// TIA Portal project "PolyMix_v0.1" (V14)

(* hardware
DEVICE "S7-1200 station_1"  S7-1200 Station
   slot 0: "Rack_0"  S7-1200 Rack  Rack  V1.0
   slot 1: "PLC_PolyMix_001"  CPU 1214C DC/DC/DC  6ES7 214-1AG40-0XB0  V4.2
DEVICE "HMI_PolyMix_001"  KTP700 Basic PN
   slot 0: "KTP700 Basic PN"  KTP700 Basic PN  6AV2 123-2GB03-0AX0  14.0.1.0
   slot 1: "HMI_RT_1"  KTP700 Basic PN  6AV2 123-2GB03-0AX0  14.0.1.0
   slot 5: "HMI_PolyMix_001.IE_CP_1"  PROFINET Interface  14.0.1.0
      slot 1: "PROFINET Interface_1"  PROFINET Interface
         slot 1: "Port_1"  Port
DEVICE "S7-1200 station_2"  S7-1200 Station
   slot 0: "Rack_0"  S7-1200 Rack  Rack  V1.0
   slot 1: "PLC_Master"  CPU 1214C DC/DC/DC  6ES7 214-1AG40-0XB0  V4.2
   slot 2: "AI 4x13BIT/AQ 2x14BIT_1"  6ES7 234-4HE32-0XB0  V2.0
   slot 3: "AI 4x13BIT/AQ 2x14BIT_2"  6ES7 234-4HE32-0XB0  V2.0
   slot 101: "CM 1241 (RS232)_1"  6ES7 241-1AH32-0XB0  V2.2
   slot 102: "CM 1241 (RS232)_2"  6ES7 241-1AH32-0XB0  V2.2
DEVICE "S7-1200 station_3"  S7-1200 Station
   slot 0: "Rack_0"  S7-1200 Rack  Rack  V1.0
   slot 1: "PLC_PolyMix_002"  CPU 1214C DC/DC/DC  6ES7 214-1AG40-0XB0  V4.2
DEVICE "HMI_PolyMix_002"  KTP700 Basic PN
   slot 0: "KTP700 Basic PN"  KTP700 Basic PN  6AV2 123-2GB03-0AX0  14.0.1.0
   slot 1: "HMI_RT_2"  KTP700 Basic PN  6AV2 123-2GB03-0AX0  14.0.1.0
   slot 5: "HMI_PolyMix_002.1.IE_CP_1"  PROFINET Interface  14.0.1.0
      slot 1: "PROFINET Interface_1"  PROFINET Interface
         slot 1: "Port_1"  Port
DEVICE "HMI_Master"  KTP700 Basic PN
   slot 0: "KTP700 Basic PN"  KTP700 Basic PN  6AV2 123-2GB03-0AX0  14.0.1.0
   slot 1: "HMI_RT_3"  KTP700 Basic PN  6AV2 123-2GB03-0AX0  14.0.1.0
   slot 5: "HMI_Master.2.1.IE_CP_1"  PROFINET Interface  14.0.1.0
      slot 1: "PROFINET Interface_1"  PROFINET Interface
         slot 1: "Port_1"  Port
DEVICE "HMI_Master_1"  KTP700 Basic PN
   slot 0: "KTP700 Basic PN"  KTP700 Basic PN  6AV2 123-2GB03-0AX0  14.0.1.0
   slot 1: "HMI_RT_4"  KTP700 Basic PN  6AV2 123-2GB03-0AX0  14.0.1.0
   slot 5: "HMI_Master.2.1.IE_CP_1"  PROFINET Interface  14.0.1.0
      slot 1: "PROFINET Interface_1"  PROFINET Interface
         slot 1: "Port_1"  Port
*)

// ===== PLC "PLC_PolyMix_001"  CPU 1214C DC/DC/DC =====
// protected blocks, not shown: "AI_ex", "AIx", "AO_ex", "DRV_M_D", "FlowMeter", "Logick", "Motors", "PLF_FC", "Time_m", "Time_r", "Time_s"

VAR_GLOBAL   // PLC tag table "Default tag table"
   "Mix_1_Clock" AT %M10.0 : Bool;
   "Mix_2_Clock" AT %M10.1 : Bool;
   "Mix_3_Clock" AT %M10.2 : Bool;
   "Flow" AT %IW256 : Int;
   "Level" AT %IW258 : Int;
END_VAR

VAR_GLOBAL   // PLC tag table "Sys"
   "pulse_01s" AT %M2.0 : Bool;
   "pulse_05s" AT %M2.1 : Bool;
   "pulse_1s" AT %M2.2 : Bool;
   "All_block" AT %M3.0 : Bool;
   "Reset_All" AT %M3.1 : Bool;
   "Sim_All" AT %M3.2 : Bool;
   "Any_Hand" AT %M5.0 : Bool;
   "DI_Hand" AT %M5.1 : Bool;
   "DO_Hand" AT %M5.2 : Bool;
   "AI_Hand" AT %M5.3 : Bool;
   "AO_Hand" AT %M5.4 : Bool;
   "M_Hand" AT %M5.5 : Bool;
   "V_Hand" AT %M5.6 : Bool;
   "X_Hand" AT %M5.7 : Bool;
   "System_Byte" AT %MB1 : Byte;
   "FirstScan" AT %M1.0 : Bool;
   "DiagStatusUpdate" AT %M1.1 : Bool;
   "ON" AT %M1.2 : Bool;
   "OFF" AT %M1.3 : Bool;
   "Clock_Byte" AT %MB0 : Byte;
   "Clock_10Hz" AT %M0.0 : Bool;
   "Clock_5Hz" AT %M0.1 : Bool;
   "Clock_2.5Hz" AT %M0.2 : Bool;
   "Clock_2Hz" AT %M0.3 : Bool;
   "Clock_1.25Hz" AT %M0.4 : Bool;
   "Clock_1Hz" AT %M0.5 : Bool;
   "Clock_0.625Hz" AT %M0.6 : Bool;
   "Clock_0.5Hz" AT %M0.7 : Bool;
   "F_pulse_01s" AT %M2.3 : Bool;
   "F_pulse_05s" AT %M2.4 : Bool;
   "F_pulse_1s" AT %M2.5 : Bool;
   "FN_pulse_01s" AT %M2.6 : Bool;
   "Clock_5s" AT %M2.7 : Bool;
   "Any_Alm" AT %M6.0 : Bool;
   "AI_Alm" AT %M6.1 : Bool;
   "M_Alm" AT %M6.2 : Bool;
   "V_Alm" AT %M6.3 : Bool;
   "C_Alm" AT %M6.4 : Bool;
   "N_Alm" AT %M6.5 : Bool;
   "L_Alm" AT %M6.6 : Bool;
   "X_Alm" AT %M6.7 : Bool;
END_VAR

VAR_GLOBAL   // PLC tag table "IO Table"
   "DD_FB_Ready" AT %I0.6 : Bool;   // I 0.6 - Дозатор сухого вещества - готовность
   "Dos_FB_Run" AT %I0.7 : Bool;   // I 0.7 - Дозатор - работа
   "DD_LLS" AT %I1.0 : Bool;   // I 1.0 - Дозатор сухого вещества - низкий уровень
   "Vibro_FB_Ready" AT %I1.1 : Bool;   // I 1.1 - Вибратор - готовность
   "Transporter" AT %I1.2 : Bool;   // I 1.2 - Пневмотранспортёр - готовность
   "DL_FB_Ready" AT %I1.3 : Bool;   // I 1.3 - Дозатор жидкого вещества - готовность
   "Dry_Run" AT %I1.4 : Bool;   // I 1.4 - Датчик протока
   "AllBlock" AT %I1.5 : Bool;   // I 1.5 - Датчик перелива или Аварийная остановка
   "M1_FB_Ready" AT %I0.0 : Bool;   // I 0.0 - Мешалка 1 - готовность
   "M1_FB_Run" AT %I0.1 : Bool;   // I 0.1 - Мешалка 1 - работа
   "M2_FB_Ready" AT %I0.2 : Bool;   // I 0.2 - Мешалка 2 - готовность
   "M2_FB_Run" AT %I0.3 : Bool;   // I 0.3 - Мешалка 2 - работа
   "M3_FB_Ready" AT %I0.4 : Bool;   // I 0.4 - Мешалка 3 - готовность
   "M3_FB_Run" AT %I0.5 : Bool;   // I 0.5 - Мешалка 3 - работа
   "M1_CMD" AT %Q0.0 : Bool;   // Q 0.0 - Мешалка 1 - запуск
   "M2_CMD" AT %Q0.1 : Bool;   // Q 0.1 - Мешалка 2 - запуск
   "M3_CMD" AT %Q0.2 : Bool;   // Q 0.2 - Мешалка 3 - запуск
   "DD_CMD" AT %Q0.3 : Bool;   // Q 0.3 - Дозатор сухого вещества - запуск
   "Vibro_CMD" AT %Q0.4 : Bool;   // Q 0.4 - Вибратор - запуск
   "DL_CMD" AT %Q0.5 : Bool;   // Q 0.5 - Дозатор жидкого вещества - запуск
   "KC1_CMD" AT %Q0.6 : Bool;   // Q 0.6 - Соленоидный клапан КС1
   "LED_Dry_Run" AT %Q0.7 : Bool;   // Q 0.7 - LED - сухой ход
   "LED_Alarm" AT %Q1.0 : Bool;   // Q 1.0 - LED - общая авария
   "LED_Empty" AT %Q1.1 : Bool;   // Q 1.1 - LED - бункер пуст
END_VAR

DATA_BLOCK "Any_DB"   // DB3
{ S7_Optimized_Access := 'FALSE' }
VERSION : 0.1
   VAR
      Level_M : Int;
      Level_S : Int;
      Flow_M : Int;
      Flow_S : Int;
      DD_View : Bool;
      Level_View : Bool;
   END_VAR
BEGIN
END_DATA_BLOCK

DATA_BLOCK "CONFIG"   // DB10
{ S7_Optimized_Access := 'FALSE' }
VERSION : 0.1
   VAR
      Config : Struct
         Use_DD : Bool;   // Использовать сухой дозатор
         Use_DL : Bool := true;   // Использовать жидкий дозатор
         Use_Mix_1 : Bool := true;   // Использовать мешалку 1
         Use_Mix_2 : Bool := true;   // Использовать мешалку 2
         Use_Mix_3 : Bool := true;   // Использовать мешалку 3
      END_STRUCT;
   END_VAR
BEGIN
END_DATA_BLOCK

DATA_BLOCK "Comm_DB"   // DB11
{ S7_Optimized_Access := 'FALSE' }
VERSION : 0.1
   VAR
      DD_Status : Int;
      DD_Mode : Int;
      DD_Alarm : Word;
      DL_Status : Int;
      DL_Mode : Int;
      DL_Alarm : Word;
      Mix_1_Status : Int;
      Mix_1_Mode : Int;
      Mix_1_Alarm : Word;
      Mix_2_Status : Int;
      Mix_2_Mode : Int;
      Mix_2_Alarm : Word;
      Mix_3_Status : Int;
      Mix_3_Mode : Int;
      Mix_3_Alarm : Word;
      KC1_Status : Int;
      Flowmeter : Real;
      Flow_Alarm : Word;
      Level : Real;
      Level_Alarm : Word;
      SP : Real;
      Start : Bool;
      Hand : Bool;
      Warning : Bool;
      Config : Struct
         Use_DD : Bool;   // Использовать сухой дозатор
         Use_DL : Bool;   // Использовать жидкий дозатор
         Use_Mix_1 : Bool;   // Использовать мешалку 1
         Use_Mix_2 : Bool;   // Использовать мешалку 2
         Use_Mix_3 : Bool;   // Использовать мешалку 3
      END_STRUCT;
      Alarm : Word;
   END_VAR
BEGIN
END_DATA_BLOCK

// folder: Modules

DATA_BLOCK "DIx_DB"   // DB200
{ S7_Optimized_Access := 'FALSE' }
VERSION : 0.1
// stored: InstanceOfName DIx
"DIx"
BEGIN
END_DATA_BLOCK

DATA_BLOCK "DOx_DB"   // DB201
{ S7_Optimized_Access := 'FALSE' }
VERSION : 0.1
// stored: InstanceOfName DOx
"DOx"
BEGIN
END_DATA_BLOCK

DATA_BLOCK "Micro_DB"   // DB207
{ S7_Optimized_Access := 'FALSE' }
VERSION : 0.1
// stored: InstanceOfName Micro
"Micro"
BEGIN
END_DATA_BLOCK

// folder: System blocks/Program resources

DATA_BLOCK "T_Reset"   // DB7
{ S7_Optimized_Access := 'TRUE' }
AUTHOR : Simatic
FAMILY : IEC
NAME : IEC_TMR
VERSION : 1.0
// stored: InstanceOfName IEC_TIMER
"IEC_TIMER"
BEGIN
END_DATA_BLOCK

DATA_BLOCK "clock_5s_ON"   // DB507
{ S7_Optimized_Access := 'TRUE' }
AUTHOR : Simatic
FAMILY : IEC
NAME : IEC_TMR
VERSION : 1.0
// stored: InstanceOfName IEC_TIMER
"IEC_TIMER"
BEGIN
END_DATA_BLOCK

DATA_BLOCK "clock_5s_OFF"   // DB508
{ S7_Optimized_Access := 'TRUE' }
AUTHOR : Simatic
FAMILY : IEC
NAME : IEC_TMR
VERSION : 1.0
// stored: InstanceOfName IEC_TIMER
"IEC_TIMER"
BEGIN
END_DATA_BLOCK

// folder: (top level)

FUNCTION "Comm_FC" : Void   // FC1, LAD
{ S7_Optimized_Access := 'TRUE' }
VERSION : 0.1
BEGIN

REGION Network 1: Сухой дозатор
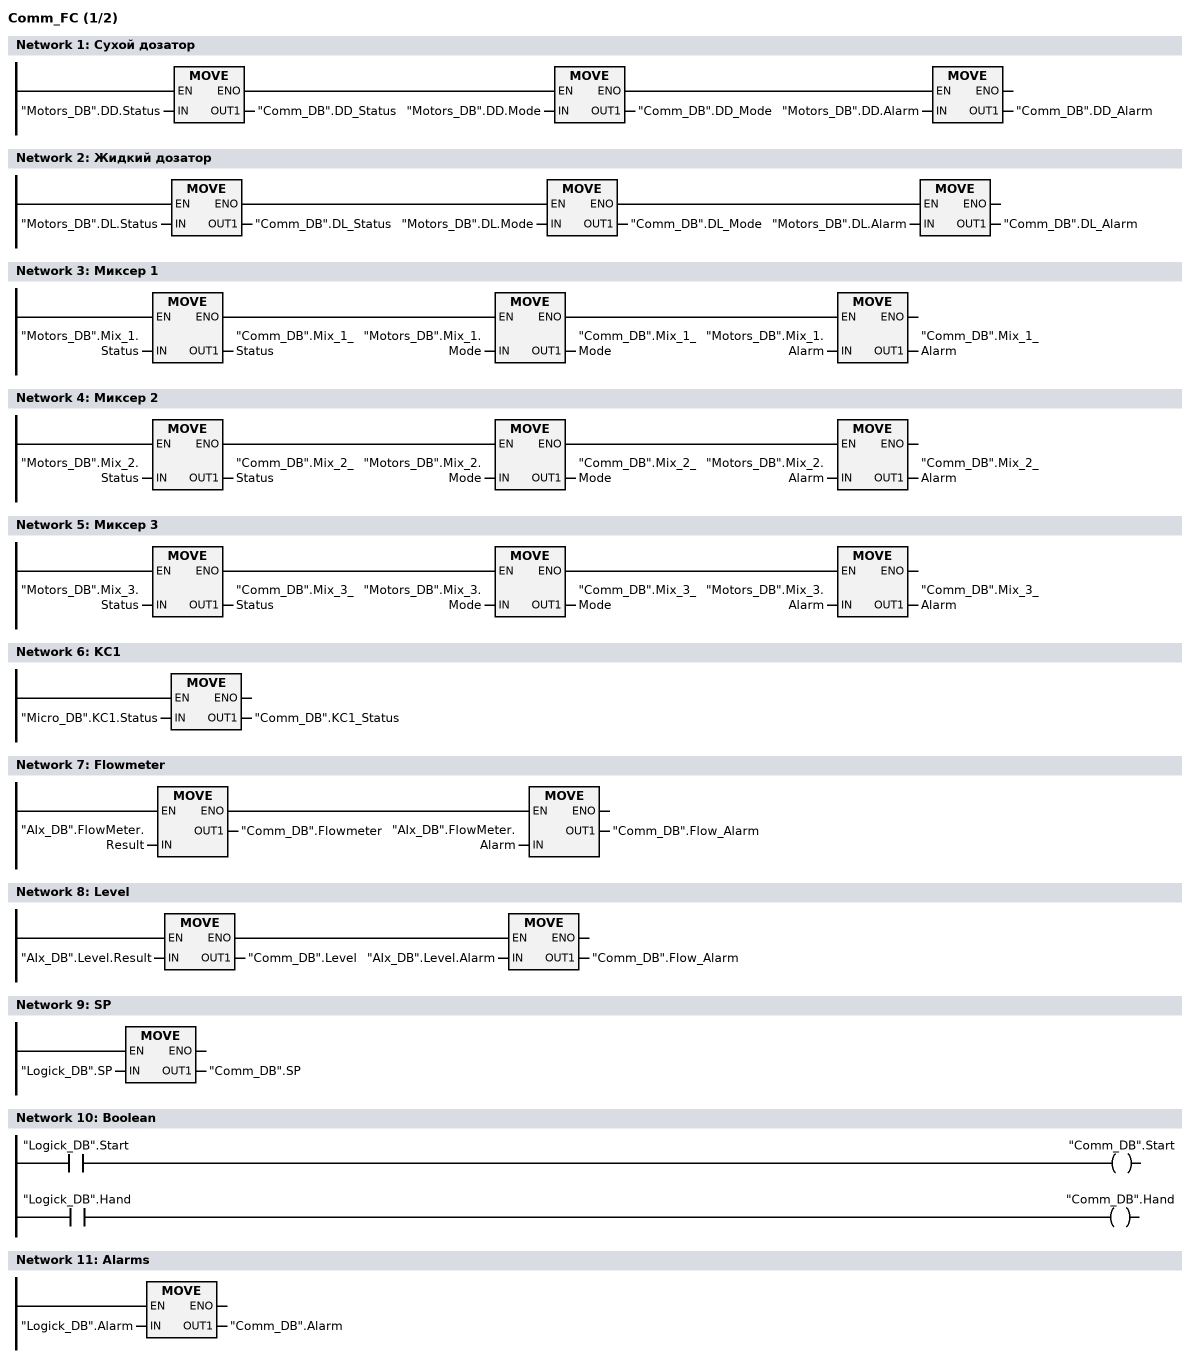
   RUNG wire#powerrail
      Move(in := "Motors_DB".DD.Status, out1 => "Comm_DB".DD_Status)
      Move(in := "Motors_DB".DD.Mode, out1 => "Comm_DB".DD_Mode)
      Move(in := "Motors_DB".DD.Alarm, out1 => "Comm_DB".DD_Alarm)
   END_RUNG
   // the same network as SCL:
   "Comm_DB".DD_Status := "Motors_DB".DD.Status;
   "Comm_DB".DD_Mode := "Motors_DB".DD.Mode;
   "Comm_DB".DD_Alarm := "Motors_DB".DD.Alarm;
END_REGION

REGION Network 2: Жидкий дозатор
   RUNG wire#powerrail
      Move(in := "Motors_DB".DL.Status, out1 => "Comm_DB".DL_Status)
      Move(in := "Motors_DB".DL.Mode, out1 => "Comm_DB".DL_Mode)
      Move(in := "Motors_DB".DL.Alarm, out1 => "Comm_DB".DL_Alarm)
   END_RUNG
   // the same network as SCL:
   "Comm_DB".DL_Status := "Motors_DB".DL.Status;
   "Comm_DB".DL_Mode := "Motors_DB".DL.Mode;
   "Comm_DB".DL_Alarm := "Motors_DB".DL.Alarm;
END_REGION

REGION Network 3: Миксер 1
   RUNG wire#powerrail
      Move(in := "Motors_DB".Mix_1.Status, out1 => "Comm_DB".Mix_1_Status)
      Move(in := "Motors_DB".Mix_1.Mode, out1 => "Comm_DB".Mix_1_Mode)
      Move(in := "Motors_DB".Mix_1.Alarm, out1 => "Comm_DB".Mix_1_Alarm)
   END_RUNG
   // the same network as SCL:
   "Comm_DB".Mix_1_Status := "Motors_DB".Mix_1.Status;
   "Comm_DB".Mix_1_Mode := "Motors_DB".Mix_1.Mode;
   "Comm_DB".Mix_1_Alarm := "Motors_DB".Mix_1.Alarm;
END_REGION

REGION Network 4: Миксер 2
   RUNG wire#powerrail
      Move(in := "Motors_DB".Mix_2.Status, out1 => "Comm_DB".Mix_2_Status)
      Move(in := "Motors_DB".Mix_2.Mode, out1 => "Comm_DB".Mix_2_Mode)
      Move(in := "Motors_DB".Mix_2.Alarm, out1 => "Comm_DB".Mix_2_Alarm)
   END_RUNG
   // the same network as SCL:
   "Comm_DB".Mix_2_Status := "Motors_DB".Mix_2.Status;
   "Comm_DB".Mix_2_Mode := "Motors_DB".Mix_2.Mode;
   "Comm_DB".Mix_2_Alarm := "Motors_DB".Mix_2.Alarm;
END_REGION

REGION Network 5: Миксер 3
   RUNG wire#powerrail
      Move(in := "Motors_DB".Mix_3.Status, out1 => "Comm_DB".Mix_3_Status)
      Move(in := "Motors_DB".Mix_3.Mode, out1 => "Comm_DB".Mix_3_Mode)
      Move(in := "Motors_DB".Mix_3.Alarm, out1 => "Comm_DB".Mix_3_Alarm)
   END_RUNG
   // the same network as SCL:
   "Comm_DB".Mix_3_Status := "Motors_DB".Mix_3.Status;
   "Comm_DB".Mix_3_Mode := "Motors_DB".Mix_3.Mode;
   "Comm_DB".Mix_3_Alarm := "Motors_DB".Mix_3.Alarm;
END_REGION

REGION Network 6: KC1
   RUNG wire#powerrail
      Move(in := "Micro_DB".KC1.Status, out1 => "Comm_DB".KC1_Status)
   END_RUNG
   // the same network as SCL:
   "Comm_DB".KC1_Status := "Micro_DB".KC1.Status;
END_REGION

REGION Network 7: Flowmeter
   RUNG wire#powerrail
      Move(in := "AIx_DB".FlowMeter.Result, out1 => "Comm_DB".Flowmeter)
      Move(in := "AIx_DB".FlowMeter.Alarm, out1 => "Comm_DB".Flow_Alarm)
   END_RUNG
   // the same network as SCL:
   "Comm_DB".Flowmeter := "AIx_DB".FlowMeter.Result;
   "Comm_DB".Flow_Alarm := "AIx_DB".FlowMeter.Alarm;
END_REGION

REGION Network 8: Level
   RUNG wire#powerrail
      Move(in := "AIx_DB".Level.Result, out1 => "Comm_DB".Level)
      Move(in := "AIx_DB".Level.Alarm, out1 => "Comm_DB".Flow_Alarm)
   END_RUNG
   // the same network as SCL:
   "Comm_DB".Level := "AIx_DB".Level.Result;
   "Comm_DB".Flow_Alarm := "AIx_DB".Level.Alarm;
END_REGION

REGION Network 9: SP
   RUNG wire#powerrail
      Move(in := "Logick_DB".SP, out1 => "Comm_DB".SP)
   END_RUNG
   // the same network as SCL:
   "Comm_DB".SP := "Logick_DB".SP;
END_REGION

REGION Network 10: Boolean
   RUNG wire#powerrail
      Contact( "Logick_DB".Start )
      Coil( "Comm_DB".Start )
   END_RUNG
   RUNG wire#powerrail
      Contact( "Logick_DB".Hand )
      Coil( "Comm_DB".Hand )
   END_RUNG
   // the same network as SCL:
   "Comm_DB".Start := "Logick_DB".Start;
   "Comm_DB".Hand := "Logick_DB".Hand;
END_REGION

REGION Network 11: Alarms
   RUNG wire#powerrail
      Move(in := "Logick_DB".Alarm, out1 => "Comm_DB".Alarm)
   END_RUNG
   // the same network as SCL:
   "Comm_DB".Alarm := "Logick_DB".Alarm;
END_REGION

REGION Network 12: Config
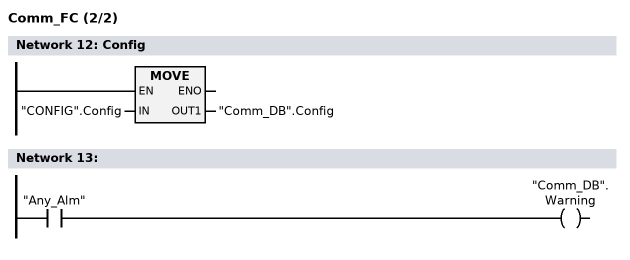
   RUNG wire#powerrail
      Move(in := "CONFIG".Config, out1 => "Comm_DB".Config)
   END_RUNG
   // the same network as SCL:
   "Comm_DB".Config := "CONFIG".Config;
END_REGION

REGION Network 13
   RUNG wire#powerrail
      Contact( "Any_Alm" )
      Coil( "Comm_DB".Warning )
   END_RUNG
   // the same network as SCL:
   "Comm_DB".Warning := "Any_Alm";
END_REGION
END_FUNCTION

ORGANIZATION_BLOCK "Main"   // OB1, LAD, ProgramCycle
TITLE = "Main Program Sweep (Cycle)"
{ S7_Optimized_Access := 'TRUE' }
VERSION : 0.1
   VAR_INPUT
      Initial_Call : Bool;   // Initial call of this OB
      Remanence : Bool;   // =True, if remanent data are available
   END_VAR
   VAR_TEMP   // added for the SCL form of the ladder/FBD networks
      _w1 : Bool;
   END_VAR
BEGIN

REGION Network 1
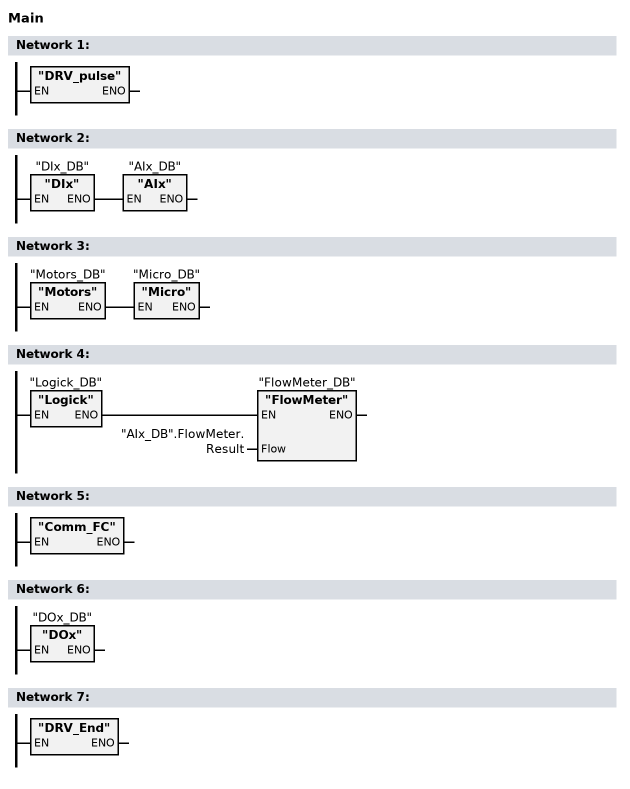
   RUNG wire#powerrail
      "DRV_pulse"()
   END_RUNG
   // the same network as SCL:
   "DRV_pulse"();
END_REGION

REGION Network 2
   RUNG wire#powerrail
      "DIx_DB"()
      "AIx_DB"()
   END_RUNG
   // the same network as SCL:
   "DIx_DB"(ENO => #_w1);   // "DIx"
   IF #_w1 THEN
       "AIx_DB"();   // "AIx"
   END_IF;
END_REGION

REGION Network 3
   RUNG wire#powerrail
      "Motors_DB"()
      "Micro_DB"()
   END_RUNG
   // the same network as SCL:
   "Motors_DB"(ENO => #_w1);   // "Motors"
   IF #_w1 THEN
       "Micro_DB"();   // "Micro"
   END_IF;
END_REGION

REGION Network 4
   RUNG wire#powerrail
      "Logick_DB"()
      "FlowMeter_DB"(Flow := "AIx_DB".FlowMeter.Result)
   END_RUNG
   // the same network as SCL:
   "Logick_DB"(ENO => #_w1);   // "Logick"
   IF #_w1 THEN
       "FlowMeter_DB"(Flow := "AIx_DB".FlowMeter.Result);   // "FlowMeter"
   END_IF;
END_REGION

REGION Network 5
   RUNG wire#powerrail
      "Comm_FC"()
   END_RUNG
   // the same network as SCL:
   "Comm_FC"();
END_REGION

REGION Network 6
   RUNG wire#powerrail
      "DOx_DB"()
   END_RUNG
   // the same network as SCL:
   "DOx_DB"();   // "DOx"
END_REGION

REGION Network 7
   RUNG wire#powerrail
      "DRV_End"()
   END_RUNG
   // the same network as SCL:
   "DRV_End"();
END_REGION
END_ORGANIZATION_BLOCK

ORGANIZATION_BLOCK "Time error interrupt"   // OB80, LAD, TimeErrorInterrupt
{ S7_Optimized_Access := 'TRUE' }
VERSION : 0.1
   VAR_INPUT
      Fault_ID : Byte;   // Fault identifier
      Csg_OBnr : OB_Any;   // Number of OB causing the error
      Csg_Prio : UInt;   // Priority of OB causing the error
   END_VAR
BEGIN
END_ORGANIZATION_BLOCK

ORGANIZATION_BLOCK "Diagnostic error interrupt"   // OB82, LAD, DiagnosticErrorInterrupt
{ S7_Optimized_Access := 'TRUE' }
VERSION : 0.1
   VAR_INPUT
      IO_State : Word;   // IO state of the HW object
      LADDR : Hw_Any;   // Hardware identifier
      Channel : UInt;   // Channel number
      MultiError : Bool;   // =true if more than one error is present
   END_VAR
BEGIN
END_ORGANIZATION_BLOCK

ORGANIZATION_BLOCK "Startup"   // OB100, LAD, Startup
TITLE = "Complete Restart"
{ S7_Optimized_Access := 'TRUE' }
VERSION : 0.1
   VAR_INPUT
      LostRetentive : Bool;   // True if retentive data are lost
      LostRTC : Bool;   // True if date and time are lost
   END_VAR
BEGIN

REGION Network 1: Запуск автоматики
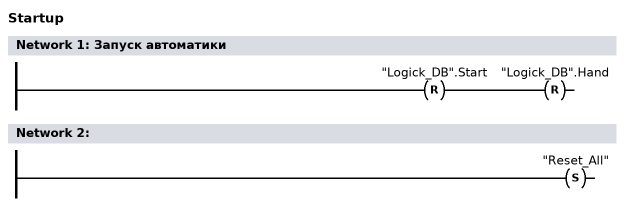
   RUNG wire#powerrail
      R_Coil( "Logick_DB".Start )
      R_Coil( "Logick_DB".Hand )
   END_RUNG
   // the same network as SCL:
   "Logick_DB".Start := FALSE;
   "Logick_DB".Hand := FALSE;
END_REGION

REGION Network 2
   RUNG wire#powerrail
      S_Coil( "Reset_All" )
   END_RUNG
   // the same network as SCL:
   "Reset_All" := TRUE;
END_REGION
END_ORGANIZATION_BLOCK

// folder: DRV_Low

FUNCTION_BLOCK "DI_ex"   // FB100, LAD
{ S7_Optimized_Access := 'FALSE' }
VERSION : 0.1
   VAR_INPUT
      Input : Bool;   // Входящий сигнал
      pulse : Bool;   // Частота фильтрации дребезка
   END_VAR
   VAR_OUTPUT
      Signal : Bool;   // Результирующий сигнал
   END_VAR
   VAR
      Hand : Bool;   // 0 - Авто, 1 - Ручной
      Start_M : Bool;   // Запуск в ручном режиме
      Data : Bool;   // Отфильтрованный сигнал
      Inverse : Bool;   // Инверсия входного сигнала
      Filter_On : Struct   // Фильтр наличия сигнала
         SP : Int;
         Now : Int;
         "Exit" : Bool;
         Start : Bool;
         Pause : Bool;
         Reset : Bool;
      END_STRUCT;
      Filter_Off : Struct   // Фильтр отсутствия сигнала
         SP : Int;
         Now : Int;
         "Exit" : Bool;
         Start : Bool;
         Pause : Bool;
         Reset : Bool;
      END_STRUCT;
      res_1 : Word;
   END_VAR
   VAR_TEMP   // added for the SCL form of the ladder/FBD networks
      _w1 : Bool;
   END_VAR
BEGIN

REGION Network 1: Устройство в ручном режиме
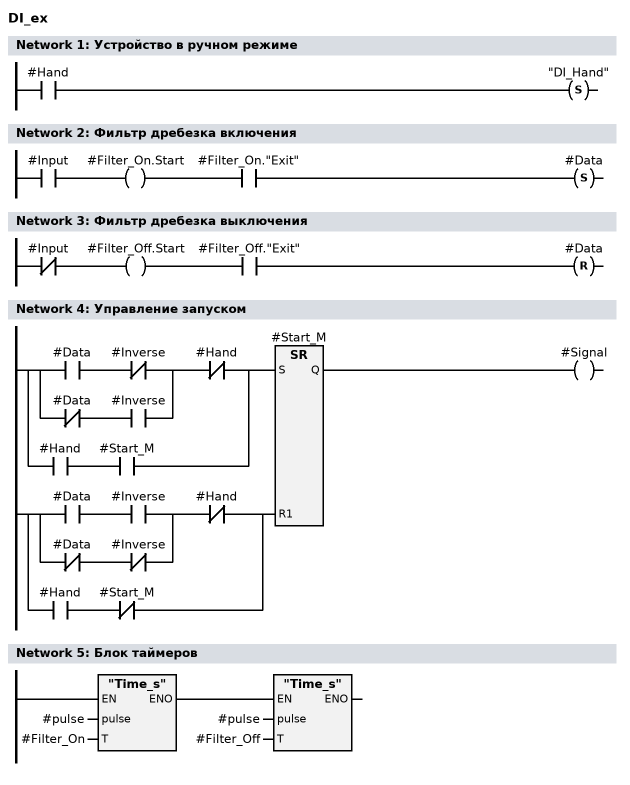
   RUNG wire#powerrail
      Contact( #Hand )
      S_Coil( "DI_Hand" )
   END_RUNG
   // the same network as SCL:
   IF #Hand THEN "DI_Hand" := TRUE; END_IF;
END_REGION

REGION Network 2: Фильтр дребезка включения
   RUNG wire#powerrail
      Contact( #Input )
      Coil( #Filter_On.Start )
      Contact( #Filter_On."Exit" )
      S_Coil( #Data )
   END_RUNG
   // the same network as SCL:
   #Filter_On.Start := #Input;
   IF #Input AND #Filter_On."Exit" THEN #Data := TRUE; END_IF;
END_REGION

REGION Network 3: Фильтр дребезка выключения
   RUNG wire#powerrail
      I_Contact( #Input )
      Coil( #Filter_Off.Start )
      Contact( #Filter_Off."Exit" )
      R_Coil( #Data )
   END_RUNG
   // the same network as SCL:
   #Filter_Off.Start := NOT #Input;
   IF NOT #Input AND #Filter_Off."Exit" THEN #Data := FALSE; END_IF;
END_REGION

REGION Network 4: Управление запуском
   RUNG wire#powerrail
      Contact( #Data )
      I_Contact( #Inverse )
      wire#w1
      I_Contact( #Hand )
      wire#w2
      S_SR(operand := #Start_M, r1 := wire#w4)
      Coil( #Signal )
   END_RUNG
   RUNG wire#powerrail
      I_Contact( #Data )
      Contact( #Inverse )
   END_RUNG wire#w1
   RUNG wire#powerrail
      Contact( #Hand )
      Contact( #Start_M )
   END_RUNG wire#w2
   RUNG wire#powerrail
      Contact( #Data )
      Contact( #Inverse )
      wire#w3
      I_Contact( #Hand )
   END_RUNG wire#w4
   RUNG wire#powerrail
      I_Contact( #Data )
      I_Contact( #Inverse )
   END_RUNG wire#w3
   RUNG wire#powerrail
      Contact( #Hand )
      I_Contact( #Start_M )
   END_RUNG wire#w4
   // the same network as SCL:
   #_w1 := (((#Data AND #Inverse) OR (NOT #Data AND NOT #Inverse)) AND NOT #Hand) OR (#Hand AND NOT #Start_M);
   IF (((#Data AND NOT #Inverse) OR (NOT #Data AND #Inverse)) AND NOT #Hand) OR (#Hand AND #Start_M) THEN
       #Start_M := TRUE;   // SR flip-flop
   END_IF;
   IF #_w1 THEN #Start_M := FALSE; END_IF;
   #Signal := #Start_M;
END_REGION

REGION Network 5: Блок таймеров
   RUNG wire#powerrail
      "Time_s"(pulse := #pulse, T := #Filter_On)
      "Time_s"(pulse := #pulse, T := #Filter_Off)
   END_RUNG
   // the same network as SCL:
   "Time_s"(pulse := #pulse, T := #Filter_On, ENO => #_w1);
   IF #_w1 THEN "Time_s"(pulse := #pulse, T := #Filter_Off); END_IF;
END_REGION
END_FUNCTION_BLOCK

FUNCTION_BLOCK "DO_ex"   // FB101, LAD
{ S7_Optimized_Access := 'FALSE' }
VERSION : 0.1
   VAR_IN_OUT
      Start_A : Bool;   // Управляющий сигнал из программы
      pulse : Bool;   // Частота длительности импульса
      Q : Bool;   // Выходной сигнал контроллера
   END_VAR
   VAR
      Hand : Bool;   // 0 - Авто, 1 - Ручной
      Start_M : Bool;   // Запуск в ручном режиме
      Simulation : Bool;   // Режим симуляции
      Inverse : Bool;   // Инверсия выхода
      Impulse : Bool;   // Импульсный режим
      T_Impulse : Struct   // Длительность импульса
         SP : Int := 5;
         Now : Int;
         "Exit" : Bool;
         Start : Bool;
         Pause : Bool;
         Reset : Bool;
      END_STRUCT;
   END_VAR
   VAR_TEMP   // added for the SCL form of the ladder/FBD networks
      _w1 : Bool;
   END_VAR
BEGIN

REGION Network 1: Устройство в ручном режиме
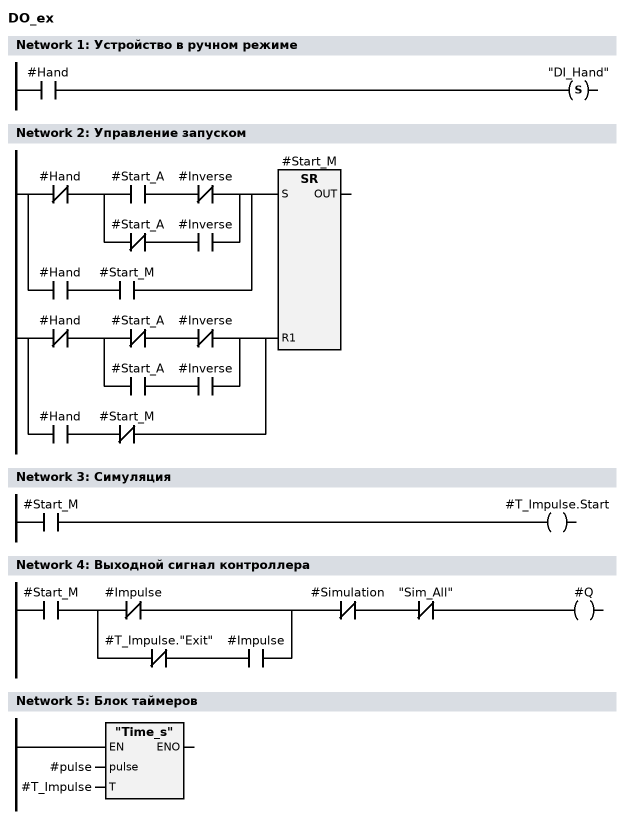
   RUNG wire#powerrail
      Contact( #Hand )
      S_Coil( "DI_Hand" )
   END_RUNG
   // the same network as SCL:
   IF #Hand THEN "DI_Hand" := TRUE; END_IF;
END_REGION

REGION Network 2: Управление запуском
   RUNG wire#powerrail
      I_Contact( #Hand )
      wire#w1
      Contact( #Start_A )
      I_Contact( #Inverse )
      wire#w2
      S_SR(operand := #Start_M, r1 := wire#w4)
   END_RUNG
   RUNG wire#w1
      I_Contact( #Start_A )
      Contact( #Inverse )
   END_RUNG wire#w2
   RUNG wire#powerrail
      Contact( #Hand )
      Contact( #Start_M )
   END_RUNG wire#w2
   RUNG wire#powerrail
      I_Contact( #Hand )
      wire#w3
      I_Contact( #Start_A )
      I_Contact( #Inverse )
   END_RUNG wire#w4
   RUNG wire#w3
      Contact( #Start_A )
      Contact( #Inverse )
   END_RUNG wire#w4
   RUNG wire#powerrail
      Contact( #Hand )
      I_Contact( #Start_M )
   END_RUNG wire#w4
   // the same network as SCL:
   #_w1 := (NOT #Hand AND ((NOT #Start_A AND NOT #Inverse) OR (#Start_A AND #Inverse))) OR (#Hand AND NOT #Start_M);
   IF (NOT #Hand AND ((#Start_A AND NOT #Inverse) OR (NOT #Start_A AND #Inverse))) OR (#Hand AND #Start_M) THEN
       #Start_M := TRUE;   // SR flip-flop
   END_IF;
   IF #_w1 THEN #Start_M := FALSE; END_IF;
END_REGION

REGION Network 3: Симуляция
   RUNG wire#powerrail
      Contact( #Start_M )
      Coil( #T_Impulse.Start )
   END_RUNG
   // the same network as SCL:
   #T_Impulse.Start := #Start_M;
END_REGION

REGION Network 4: Выходной сигнал контроллера
   RUNG wire#powerrail
      Contact( #Start_M )
      wire#w1
      I_Contact( #Impulse )
      wire#w2
      I_Contact( #Simulation )
      I_Contact( "Sim_All" )
      Coil( #Q )
   END_RUNG
   RUNG wire#w1
      I_Contact( #T_Impulse."Exit" )
      Contact( #Impulse )
   END_RUNG wire#w2
   // the same network as SCL:
   #Q := #Start_M AND (NOT #Impulse OR (NOT #T_Impulse."Exit" AND #Impulse)) AND NOT #Simulation AND NOT "Sim_All";
END_REGION

REGION Network 5: Блок таймеров
   RUNG wire#powerrail
      "Time_s"(pulse := #pulse, T := #T_Impulse)
   END_RUNG
   // the same network as SCL:
   "Time_s"(pulse := #pulse, T := #T_Impulse);
END_REGION
END_FUNCTION_BLOCK

FUNCTION_BLOCK "DRV_Micro"   // FB104, LAD
{ S7_Optimized_Access := 'FALSE' }
VERSION : 0.1
   VAR_INPUT
      Start_A : Bool;   // Запрос запуска
      FB : Bool;   // ОС
      Reset : Bool;   // Сброс аварий
      All_Block : Bool;   // Блокировка
   END_VAR
   VAR_OUTPUT
      CMD : Bool;   // Команда
   END_VAR
   VAR_IN_OUT
      Alarm : Bool;   // Авария
   END_VAR
   VAR
      Hand : Bool;   // Ручной режим
      Start_M : Bool;   // Запуск в ручном режиме
      No_FB : Bool;   // Не использовать ОС
      ON : Bool;   // Успешно запущено
      OFF : Bool;   // Успешно остановлено
      Status : Int;   // Статус устройства / Статус привода
      Wait_On : Struct   // Ожидание ОС контактора / Время на запуск
         SP : Int := 2;
         Now : Int;
         "Exit" : Bool;
         Start : Bool;
         Pause : Bool;
         Reset : Bool;
      END_STRUCT;
      Wait_Off : Struct   // Ожидание концевиков / Время на останов
         SP : Int := 2;
         Now : Int;
         "Exit" : Bool;
         Start : Bool;
         Pause : Bool;
         Reset : Bool;
      END_STRUCT;
   END_VAR
   VAR_TEMP   // added for the SCL form of the ladder/FBD networks
      _w1 : Bool;
      _w2 : Bool;
   END_VAR
BEGIN

REGION Network 1: Управление запуском / дискретный управляющий сигнал
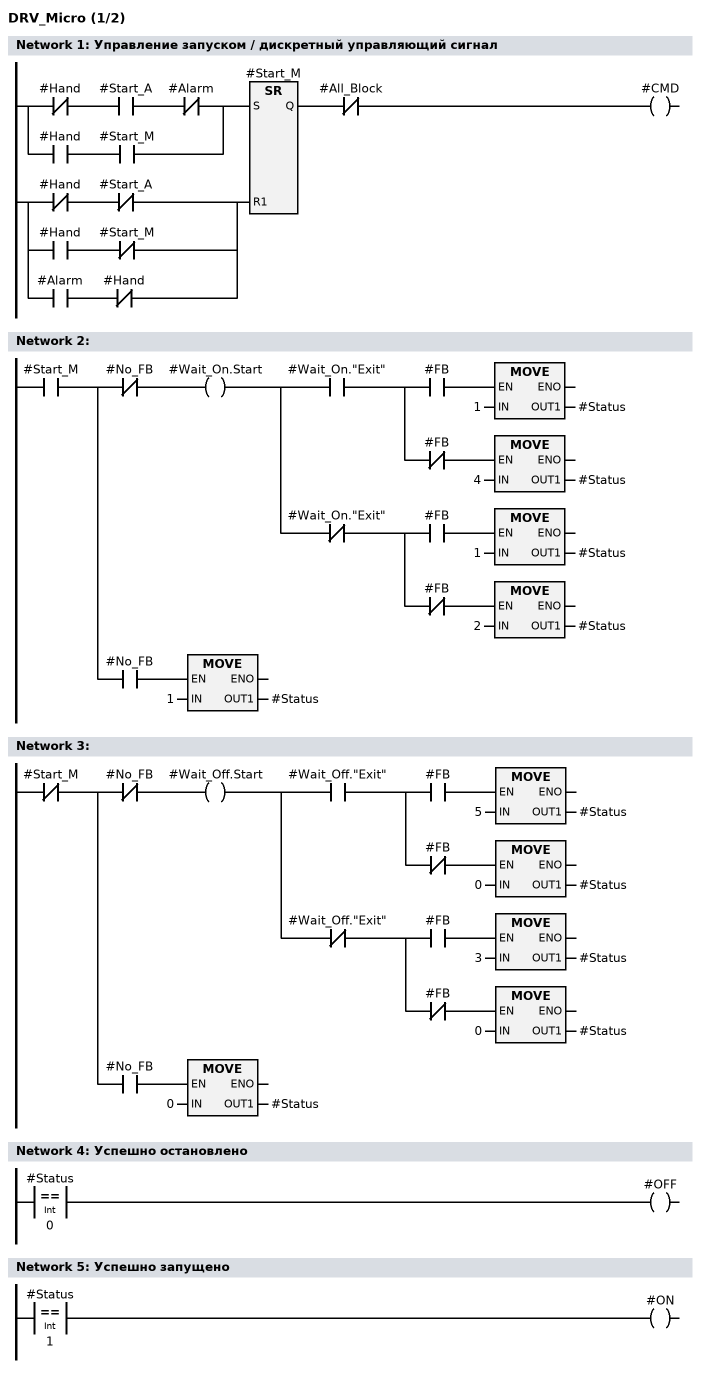
   RUNG wire#powerrail
      I_Contact( #Hand )
      Contact( #Start_A )
      I_Contact( #Alarm )
      wire#w1
      S_SR(operand := #Start_M, r1 := wire#w2)
      I_Contact( #All_Block )
      Coil( #CMD )
   END_RUNG
   RUNG wire#powerrail
      Contact( #Hand )
      Contact( #Start_M )
   END_RUNG wire#w1
   RUNG wire#powerrail
      I_Contact( #Hand )
      I_Contact( #Start_A )
   END_RUNG wire#w2
   RUNG wire#powerrail
      Contact( #Hand )
      I_Contact( #Start_M )
   END_RUNG wire#w2
   RUNG wire#powerrail
      Contact( #Alarm )
      I_Contact( #Hand )
   END_RUNG wire#w2
   // the same network as SCL:
   #_w1 := (NOT #Hand AND NOT #Start_A) OR (#Hand AND NOT #Start_M) OR (#Alarm AND NOT #Hand);
   IF (NOT #Hand AND #Start_A AND NOT #Alarm) OR (#Hand AND #Start_M) THEN
       #Start_M := TRUE;   // SR flip-flop
   END_IF;
   IF #_w1 THEN #Start_M := FALSE; END_IF;
   #CMD := #Start_M AND NOT #All_Block;
END_REGION

REGION Network 2
   RUNG wire#powerrail
      Contact( #Start_M )
      wire#w1
      I_Contact( #No_FB )
      Coil( #Wait_On.Start )
      wire#w2
      Contact( #Wait_On."Exit" )
      wire#w3
      Contact( #FB )
      Move(in := 1, out1 => #Status)
   END_RUNG
   RUNG wire#w3
      I_Contact( #FB )
      Move(in := 4, out1 => #Status)
   END_RUNG
   RUNG wire#w2
      I_Contact( #Wait_On."Exit" )
      wire#w4
      Contact( #FB )
      Move(in := 1, out1 => #Status)
   END_RUNG
   RUNG wire#w4
      I_Contact( #FB )
      Move(in := 2, out1 => #Status)
   END_RUNG
   RUNG wire#w1
      Contact( #No_FB )
      Move(in := 1, out1 => #Status)
   END_RUNG
   // the same network as SCL:
   #Wait_On.Start := #Start_M AND NOT #No_FB;
   #_w1 := #Wait_On.Start AND #Wait_On."Exit";
   IF #_w1 AND #FB THEN #Status := 1; END_IF;
   IF #_w1 AND NOT #FB THEN #Status := 4; END_IF;
   #_w2 := #Wait_On.Start AND NOT #Wait_On."Exit";
   IF #_w2 AND #FB THEN #Status := 1; END_IF;
   IF #_w2 AND NOT #FB THEN #Status := 2; END_IF;
   IF #Start_M AND #No_FB THEN #Status := 1; END_IF;
END_REGION

REGION Network 3
   RUNG wire#powerrail
      I_Contact( #Start_M )
      wire#w1
      I_Contact( #No_FB )
      Coil( #Wait_Off.Start )
      wire#w2
      Contact( #Wait_Off."Exit" )
      wire#w3
      Contact( #FB )
      Move(in := 5, out1 => #Status)
   END_RUNG
   RUNG wire#w3
      I_Contact( #FB )
      Move(in := 0, out1 => #Status)
   END_RUNG
   RUNG wire#w2
      I_Contact( #Wait_Off."Exit" )
      wire#w4
      Contact( #FB )
      Move(in := 3, out1 => #Status)
   END_RUNG
   RUNG wire#w4
      I_Contact( #FB )
      Move(in := 0, out1 => #Status)
   END_RUNG
   RUNG wire#w1
      Contact( #No_FB )
      Move(in := 0, out1 => #Status)
   END_RUNG
   // the same network as SCL:
   #Wait_Off.Start := NOT #Start_M AND NOT #No_FB;
   #_w1 := #Wait_Off.Start AND #Wait_Off."Exit";
   IF #_w1 AND #FB THEN #Status := 5; END_IF;
   IF #_w1 AND NOT #FB THEN #Status := 0; END_IF;
   #_w2 := #Wait_Off.Start AND NOT #Wait_Off."Exit";
   IF #_w2 AND #FB THEN #Status := 3; END_IF;
   IF #_w2 AND NOT #FB THEN #Status := 0; END_IF;
   IF NOT #Start_M AND #No_FB THEN #Status := 0; END_IF;
END_REGION

REGION Network 4: Успешно остановлено
   RUNG wire#powerrail
      { S7_Templates := "SrcType := Int" } EQ_Contact(in1 := #Status, in2 := 0)
      Coil( #OFF )
   END_RUNG
   // the same network as SCL:
   #OFF := #Status = 0;
END_REGION

REGION Network 5: Успешно запущено
   RUNG wire#powerrail
      { S7_Templates := "SrcType := Int" } EQ_Contact(in1 := #Status, in2 := 1)
      Coil( #ON )
   END_RUNG
   // the same network as SCL:
   #ON := #Status = 1;
END_REGION

REGION Network 6: Авария